// TIA Portal project "Mel7_new" (V15.1)

(* hardware
DEVICE "Станция S7-1200_1"  S7-1200 Station
   slot 0: "Rack_0"  S7-1200 Rack  Rack  V1.0
   slot 1: "01_CPU"  CPU 1215C DC/DC/DC  6ES7 215-1AG40-0XB0  V4.2
   slot 2: "AI 8x13 бит_1"  6ES7 231-4HF32-0XB0  V2.0
   slot 3: "AI 8x13 бит_2"  6ES7 231-4HF32-0XB0  V2.0
   slot 4: "AI 8x13 бит_3"  6ES7 231-4HF32-0XB0  V2.0
   slot 5: "AI 8x13 бит_4"  6ES7 231-4HF32-0XB0  V2.0
   slot 6: "AI 8xRTD_1"  SM 1231 AI8 x RTD  6ES7 231-5PF32-0XB0  V2.0
   slot 7: "AI 8xRTD_2"  SM 1231 AI8 x RTD  6ES7 231-5PF32-0XB0  V2.0
   slot 101: "CM 1243-5"  CM 1243-5  6GK7 243-5DX30-0XE0  V1.3
DEVICE "02_HMI"  KTP1200 Basic PN
   slot 0: "02_HMI"  KTP1200 Basic PN  6AV2 123-2MB03-0AX0  15.1.0.0
   slot 1: "HMI_RT_1"  KTP1200 Basic PN  6AV2 123-2MB03-0AX0  15.1.0.0
   slot 5: "02_HMI.IE_CP_1"  PROFINET Interface  15.0.1.0
      slot 1: "PROFINET Interface_1"  PROFINET Interface
         slot 1: "Port_1"  Port
DEVICE "S7300/ET200M station_1"  S7-300 station
   slot 0: "Rail_0"  Rail  6ES7 390-1***0-0AA0
   slot 2: "Slave_1"  IM 153-2  6ES7 153-2BA10-0XB0  V6.0
   slot 4: "DI 32x24VDC_1"  DI32 x 24VDC  6ES7 321-1BL00-0AA0
   slot 5: "DO 16x24VDC/0.5A_1"  DO16 x 24VDC / 0.5A  6ES7 322-1BH01-0AA0
   slot 6: "DO 16x24VDC/0.5A_2"  DO16 x 24VDC / 0.5A  6ES7 322-1BH01-0AA0
   slot 7: "AO 8x12BIT_1"  AO8 x 12 bits  6ES7 332-5HF00-0AB0
*)

// ===== PLC "01_CPU"  CPU 1215C DC/DC/DC =====

VAR_GLOBAL   // PLC tag table "Стандартная таблица переменных"
   "System_Byte" AT %MB1 : Byte;
   "FirstScan" AT %M1.0 : Bool;
   "DiagStatusUpdate" AT %M1.1 : Bool;
   "AlwaysTRUE" AT %M1.2 : Bool;
   "AlwaysFALSE" AT %M1.3 : Bool;
   "Clock_Byte" AT %MB0 : Byte;
   "Clock_10Hz" AT %M0.0 : Bool;
   "Clock_5Hz" AT %M0.1 : Bool;
   "Clock_2.5Hz" AT %M0.2 : Bool;
   "Clock_2Hz" AT %M0.3 : Bool;
   "Clock_1.25Hz" AT %M0.4 : Bool;
   "Clock_1Hz" AT %M0.5 : Bool;
   "Clock_0.625Hz" AT %M0.6 : Bool;
   "Clock_0.5Hz" AT %M0.7 : Bool;
END_VAR

TYPE "AI_STR"
   STRUCT
      "Кнопка: Закрыть фейсплату" : Bool;
      "Кнопка: Активировать HH" : Bool;   // Активация уставки НН
      "Кнопка: Активировать H" : Bool;   // Активация уставки Н
      "Кнопка: Активировать L" : Bool;   // Активация уставки L
      "Кнопка: Активировать LL" : Bool;   // Активация уставки LL
      "Кнопка: Ремонт" : Bool;   // Активация кнопки Ремонт
      Видимость : Bool;   // Видимость
      "Индикатор: Зашкал" : Bool;   // Overflow
      "Индикатор: Перелёт" : Bool;   // Overshoot range
      "Авария: Выход за HH" : Bool;   // Выход за уставку НН
      "Предупреждение: Выход за H" : Bool;   // Выход за уставку Н
      "Предупреждение: Выход за L" : Bool;   // Выход за уставку L
      "Авария: Выход за LL" : Bool;   // Выход за уставку LL
      "Индикатор: Недолет" : Bool;   // Undershoot range
      "Индикатор: Обрыв" : Bool;   // Underflow
      "Индикатор: В норме" : Bool;
      "Индикатор: HH активирована" : Bool;
      "Индикатор: H активирована" : Bool;
      "Индикатор: L активирована" : Bool;
      "Индикатор: LL активирована" : Bool;
      "Уставка: MAX" : Real := 100.0;   // Верхняя граница шкалы прибора
      "Уставка: MIN" : Real := 0.0;   // Нижняя граница шкалы прибора
      "Уставка: HH" : Real := 80.0;   // Верхняя аварийная уставка
      "Уставка: H" : Real := 70.0;   // Верхняя предупредительная уставка
      "Уставка: L" : Real := 15.0;   // Нижняя предупредительная уставка
      "Уставка: LL" : Real := 10.0;   // Нижняя аварийная уставка
      "Уставка: Перелёт" : Real := 20.0;   // Overshoot
      "Уставка: Недолёт" : Real := 4.0;   // Undershoot
      PV : Real;   // Переменная процесса
      Ток : Real;   // Токовый сигнал мА
      AnimCode : Int;
      Error : Word;   // Регистр функции ошибки
      Bipolar : Bool;   // 1 - биполярный сигнал, 0 - униполярный сигнал
      Overshoot_MIN : Int := 27649;
      Undershoot_MAX : Int := -1;
   END_STRUCT;
END_TYPE

TYPE "Motor_S"
VERSION : 0.1
   STRUCT
      Mode : Bool;   // Режим Оператор=0 Режим Автомат=1
      OperatorStart : Bool;   // Старт в режиме оператор
      AutoStart : Bool;
      ResetAlarm : Bool;
      ResetWorkTime : Bool;   // Сброс часов работы мотора
      AnimCode : Int;
      WorkTime : DInt;   // Время работы мотора
      TimeOutAccMotor : Int;
   END_STRUCT;
END_TYPE

TYPE "PID_CONT S"
   STRUCT
      COM_RST : Bool;   // Полный рестарт
      LMNR_HS : Bool;   // Верхняя граница сигнала позиционной обратной связи
      LMNR_LS : Bool;   // Нижняя граница сигнала позиционной обратной связи
      LMNS_ON : Bool := true;   // Включение сигнала ручного воздействия
      LMNUP : Bool;   // Увеличение управляющих сигналов
      LMNDN : Bool;   // Уменьшение управляющих сигналов
      PVPER_ON : Bool;   // Включение переменной процесса периферии
      CYCLE : Time := T#1s;   // Время опроса
      SP_INT : Real;   // Внутренне значение уставки
      PV_IN : Real;   // Ввод переменной уставки
      PV_PER : Word;   // Переменная процесса от периферии
      GAIN : Real := 2.0;   // Коэффицент пропорциональности
      TI : Time := T#20s;   // Время интегрирования
      DEADB_W : Real := 1.0;   // Ширина зоны нечувствительности
      PV_FAC : Real := 1.0;   // Коээфицент переменной процесса
      PV_OFF : Real;   // Смещение переменной процесса
      PULSE_TM : Time := T#3s;   // Минимальная длительность импульса
      BREAK_TM : Time := T#3s;   // Минимальная время пауза
      MTR_TM : Time := T#30s;   // Время прогона привода
      DISV : Real;   // Возмущающее воздействие
      QLMNUP : Bool;   // Увеличение управляющего сигнала
      QLMNDN : Bool;   // Уменьшение управляющего сигнала
      PV : Real;   // Переменная процесса
      ER : Real;   // Сигнал ошибки
   END_STRUCT;
END_TYPE

TYPE "DI_STR"
   STRUCT
      "BOOL" : Bool;
      "INT" : Int;
   END_STRUCT;
END_TYPE

TYPE "PID_STR"
VERSION : 0.1
   STRUCT
      SP : Real;
      PV : Real;
      Gain : Real := 2.0;
      Ti : Time := T#20s;
      Td : Time := T#10s;
      Tm_lag : Time := T#2s;
      Man_ON : Bool := true;
      MAN : Real;
      LMN_HI : Real := 100.0;
      LMN_LO : Real := 0.0;
      Reset : Bool;
      LMN : Real;
   END_STRUCT;
END_TYPE

TYPE "Motor_STR"
VERSION : 0.1
   STRUCT
      AnimCodeMotor : Int;   // Код анимации мотора
      AnimCodeKey : Int;   // Код анимации ключа: =0 Сблокированный,=1 Ручной =10,11-Ошибочная сигнализация
      TimeOutPreMotor : Int := 4;   // Таймер на нарушения мотора уставка
      TimeOutAccMotor : Int;   // Таймер на нарушения мотора аккомулятор
      TimeOutPreKey : Int := 2;   // Таймер на нарушение положения ключа уставка
      TimeOutACCKey : Int;   // Таймер на нарушение положения ключа аккомулятор
      Mode : Int;   // Режим Оператор=0 Режим Автомат=1
      PouseBeetwenON : Word;   // Пауза между включениями мотора
      WorkTime : DInt;   // Время работы мотора
      OperatorStart : Bool;   // Старт в режиме оператор
      ResetAlr : Bool;   // Сброс нарушений
      ResetWorkTime : Bool;   // Сброс часов работы мотора
      Start : Bool;   // Старт Мотора
      StartPulse : Bool;   // Старт Мотора пульс
      ModeBool : Bool;
   END_STRUCT;
END_TYPE

TYPE "Narabotki"
   STRUCT
      Hour : DInt;
      Minute : Int;
      Second : Int;
      old : Bool;
      reset : Bool;
   END_STRUCT;
END_TYPE

TYPE "Valve_STR"
VERSION : 0.1
   STRUCT
      AnimCodeValve : Int;   // Код анимации крана: =0 Нейтр,=1 Открыт, =3 закрыт, >10 Нарушения
      AnimCodeKey : Int;   // Код анимации ключа: =0 Сблокированный,=1 Ручной =10,11-Ошибочная сигнализация
      TimeOutPreValve : Int := 60;   // Таймер на нарушения движения уставка
      TimeOutAccValve : Int;   // Таймер на нарушения мотора аккомулятор
      TimeOutPreKey : Int := 2;   // Таймер на нарушение положения ключа уставка
      TimeOutACCKey : Int;   // Таймер на нарушение положения ключа аккомулятор
      Mode : Int;   // Режим Оператор=0 Режим Автомат=1
      PouseBeetwenON : Word := 16#0;   // Пауза между включениями мотора
      WorkTime : DInt;   // Время работы мотора
      OperatorOpen : Bool;   // Открытие в режиме опреатор
      OperatorClose : Bool;   // Закрытие в режиме опреатор
      ResetAlr : Bool;   // Сброс нарушений
      ResetWorkTime : Bool;   // Сброс часов работы крана
      CmdOpen : Bool;   // Команда на открытие
      CmdOpenPulse : Bool;   // Команда на открытие пульс
      CmdClose : Bool;   // Команда на закрытие
      CmdClosePulse : Bool;   // Команда на закрытие пульс
   END_STRUCT;
END_TYPE

DATA_BLOCK "01_DB_AI"   // DB1
{ S7_Optimized_Access := 'FALSE' }
VERSION : 0.1
   VAR
      L_1c : "AI_STR";
      L_1c_1 : "AI_STR";
      L_1c_2 : "AI_STR";
      L_1c_3 : "AI_STR";
      L_1c_4 : "AI_STR";
      L_1c_5 : "AI_STR";
      L_1c_6 : "AI_STR";
      L_1c_7 : "AI_STR";
      L_1c_8 : "AI_STR";
      L_1c_9 : "AI_STR";
      L_1c_10 : "AI_STR";
      L_1c_11 : "AI_STR";
      L_1c_12 : "AI_STR";
      L_1c_13 : "AI_STR";
      L_1c_14 : "AI_STR";
      L_1c_15 : "AI_STR";
      L_1c_16 : "AI_STR";
      L_1c_17 : "AI_STR";
      L_1c_18 : "AI_STR";
      L_1c_19 : "AI_STR";
      L_1c_20 : "AI_STR";
      L_1c_21 : "AI_STR";
      L_1c_22 : "AI_STR";
      L_1c_23 : "AI_STR";
      L_1c_24 : "AI_STR";
      L_1c_25 : "AI_STR";
      L_1c_26 : "AI_STR";
      L_1c_27 : "AI_STR";
      L_1c_28 : "AI_STR";
      L_1c_29 : "AI_STR";
      L_1c_30 : "AI_STR";
      L_1c_31 : "AI_STR";
      L_1c_32 : "AI_STR";
      L_1c_33 : "AI_STR";
      L_1c_36 : "AI_STR";
      L_1c_37 : "AI_STR";
      L_1c_38 : "AI_STR";
      L_1c_39 : "AI_STR";
      L_1c_40 : "AI_STR";
      L_1c_41 : "AI_STR";
      L_1c_42 : "AI_STR";
      L_1c_43 : "AI_STR";
      L_1c_44 : "AI_STR";
      L_1c_45 : "AI_STR";   // Расход руды tarir
   END_VAR
BEGIN
   L_1c_20."Кнопка: Активировать HH" := TRUE;
   L_1c_26."Кнопка: Активировать HH" := FALSE;
   L_1c."Кнопка: Закрыть фейсплату" := FALSE;
   L_1c."Кнопка: Активировать HH" := FALSE;
   L_1c."Кнопка: Активировать H" := FALSE;
   L_1c."Кнопка: Активировать L" := FALSE;
   L_1c."Кнопка: Активировать LL" := FALSE;
   L_1c."Кнопка: Ремонт" := FALSE;
   L_1c.Видимость := FALSE;
   L_1c."Индикатор: Зашкал" := FALSE;
   L_1c."Индикатор: Перелёт" := FALSE;
   L_1c."Авария: Выход за HH" := FALSE;
   L_1c."Предупреждение: Выход за H" := FALSE;
   L_1c."Предупреждение: Выход за L" := FALSE;
   L_1c."Авария: Выход за LL" := FALSE;
   L_1c."Индикатор: Недолет" := FALSE;
   L_1c."Индикатор: Обрыв" := FALSE;
   L_1c."Индикатор: В норме" := FALSE;
   L_1c."Индикатор: HH активирована" := FALSE;
   L_1c."Индикатор: H активирована" := FALSE;
   L_1c."Индикатор: L активирована" := FALSE;
   L_1c."Индикатор: LL активирована" := FALSE;
   L_1c."Уставка: MAX" := 100.0;
   L_1c."Уставка: MIN" := 0.0;
   L_1c."Уставка: HH" := 80.0;
   L_1c."Уставка: H" := 70.0;
   L_1c."Уставка: L" := 15.0;
   L_1c."Уставка: LL" := 10.0;
   L_1c."Уставка: Перелёт" := 20.0;
   L_1c."Уставка: Недолёт" := 4.0;
   L_1c.PV := 3.204572;
   L_1c.Ток := 4.512732;
   L_1c.AnimCode := 0;
   L_1c.Error := 16#0000;
   L_1c.Bipolar := FALSE;
   L_1c.Overshoot_MIN := 27649;
   L_1c.Undershoot_MAX := -1;
   L_1c_1."Кнопка: Закрыть фейсплату" := FALSE;
   L_1c_1."Кнопка: Активировать HH" := FALSE;
   L_1c_1."Кнопка: Активировать H" := FALSE;
   L_1c_1."Кнопка: Активировать L" := FALSE;
   L_1c_1."Кнопка: Активировать LL" := FALSE;
   L_1c_1."Кнопка: Ремонт" := FALSE;
   L_1c_1.Видимость := FALSE;
   L_1c_1."Индикатор: Зашкал" := FALSE;
   L_1c_1."Индикатор: Перелёт" := FALSE;
   L_1c_1."Авария: Выход за HH" := FALSE;
   L_1c_1."Предупреждение: Выход за H" := FALSE;
   L_1c_1."Предупреждение: Выход за L" := FALSE;
   L_1c_1."Авария: Выход за LL" := FALSE;
   L_1c_1."Индикатор: Недолет" := FALSE;
   L_1c_1."Индикатор: Обрыв" := FALSE;
   L_1c_1."Индикатор: В норме" := FALSE;
   L_1c_1."Индикатор: HH активирована" := FALSE;
   L_1c_1."Индикатор: H активирована" := FALSE;
   L_1c_1."Индикатор: L активирована" := FALSE;
   L_1c_1."Индикатор: LL активирована" := FALSE;
   L_1c_1."Уставка: MAX" := 100.0;
   L_1c_1."Уставка: MIN" := 0.0;
   L_1c_1."Уставка: HH" := 80.0;
   L_1c_1."Уставка: H" := 70.0;
   L_1c_1."Уставка: L" := 15.0;
   L_1c_1."Уставка: LL" := 10.0;
   L_1c_1."Уставка: Перелёт" := 20.0;
   L_1c_1."Уставка: Недолёт" := 4.0;
   L_1c_1.PV := 13.17636;
   L_1c_1.Ток := 6.108218;
   L_1c_1.AnimCode := 0;
   L_1c_1.Error := 16#0000;
   L_1c_1.Bipolar := FALSE;
   L_1c_1.Overshoot_MIN := 27649;
   L_1c_1.Undershoot_MAX := -1;
   L_1c_2."Кнопка: Закрыть фейсплату" := FALSE;
   L_1c_2."Кнопка: Активировать HH" := FALSE;
   L_1c_2."Кнопка: Активировать H" := FALSE;
   L_1c_2."Кнопка: Активировать L" := FALSE;
   L_1c_2."Кнопка: Активировать LL" := FALSE;
   L_1c_2."Кнопка: Ремонт" := FALSE;
   L_1c_2.Видимость := FALSE;
   L_1c_2."Индикатор: Зашкал" := FALSE;
   L_1c_2."Индикатор: Перелёт" := FALSE;
   L_1c_2."Авария: Выход за HH" := FALSE;
   L_1c_2."Предупреждение: Выход за H" := FALSE;
   L_1c_2."Предупреждение: Выход за L" := FALSE;
   L_1c_2."Авария: Выход за LL" := FALSE;
   L_1c_2."Индикатор: Недолет" := FALSE;
   L_1c_2."Индикатор: Обрыв" := FALSE;
   L_1c_2."Индикатор: В норме" := FALSE;
   L_1c_2."Индикатор: HH активирована" := FALSE;
   L_1c_2."Индикатор: H активирована" := FALSE;
   L_1c_2."Индикатор: L активирована" := FALSE;
   L_1c_2."Индикатор: LL активирована" := FALSE;
   L_1c_2."Уставка: MAX" := 100.0;
   L_1c_2."Уставка: MIN" := 0.0;
   L_1c_2."Уставка: HH" := 90.0;
   L_1c_2."Уставка: H" := 70.0;
   L_1c_2."Уставка: L" := 15.0;
   L_1c_2."Уставка: LL" := 10.0;
   L_1c_2."Уставка: Перелёт" := 20.0;
   L_1c_2."Уставка: Недолёт" := 4.0;
   L_1c_2.PV := 69.30339;
   L_1c_2.Ток := 15.08854;
   L_1c_2.AnimCode := 0;
   L_1c_2.Error := 16#0000;
   L_1c_2.Bipolar := FALSE;
   L_1c_2.Overshoot_MIN := 27649;
   L_1c_2.Undershoot_MAX := -1;
   L_1c_3."Кнопка: Закрыть фейсплату" := FALSE;
   L_1c_3."Кнопка: Активировать HH" := FALSE;
   L_1c_3."Кнопка: Активировать H" := FALSE;
   L_1c_3."Кнопка: Активировать L" := FALSE;
   L_1c_3."Кнопка: Активировать LL" := FALSE;
   L_1c_3."Кнопка: Ремонт" := FALSE;
   L_1c_3.Видимость := FALSE;
   L_1c_3."Индикатор: Зашкал" := FALSE;
   L_1c_3."Индикатор: Перелёт" := FALSE;
   L_1c_3."Авария: Выход за HH" := FALSE;
   L_1c_3."Предупреждение: Выход за H" := FALSE;
   L_1c_3."Предупреждение: Выход за L" := FALSE;
   L_1c_3."Авария: Выход за LL" := FALSE;
   L_1c_3."Индикатор: Недолет" := FALSE;
   L_1c_3."Индикатор: Обрыв" := FALSE;
   L_1c_3."Индикатор: В норме" := FALSE;
   L_1c_3."Индикатор: HH активирована" := FALSE;
   L_1c_3."Индикатор: H активирована" := FALSE;
   L_1c_3."Индикатор: L активирована" := FALSE;
   L_1c_3."Индикатор: LL активирована" := FALSE;
   L_1c_3."Уставка: MAX" := 100.0;
   L_1c_3."Уставка: MIN" := 0.0;
   L_1c_3."Уставка: HH" := 80.0;
   L_1c_3."Уставка: H" := 70.0;
   L_1c_3."Уставка: L" := 15.0;
   L_1c_3."Уставка: LL" := 10.0;
   L_1c_3."Уставка: Перелёт" := 20.0;
   L_1c_3."Уставка: Недолёт" := 4.0;
   L_1c_3.PV := 7.895689;
   L_1c_3.Ток := 5.26331;
   L_1c_3.AnimCode := 0;
   L_1c_3.Error := 16#0000;
   L_1c_3.Bipolar := FALSE;
   L_1c_3.Overshoot_MIN := 27649;
   L_1c_3.Undershoot_MAX := -1;
   L_1c_4."Кнопка: Закрыть фейсплату" := FALSE;
   L_1c_4."Кнопка: Активировать HH" := FALSE;
   L_1c_4."Кнопка: Активировать H" := FALSE;
   L_1c_4."Кнопка: Активировать L" := FALSE;
   L_1c_4."Кнопка: Активировать LL" := FALSE;
   L_1c_4."Кнопка: Ремонт" := FALSE;
   L_1c_4.Видимость := FALSE;
   L_1c_4."Индикатор: Зашкал" := FALSE;
   L_1c_4."Индикатор: Перелёт" := FALSE;
   L_1c_4."Авария: Выход за HH" := FALSE;
   L_1c_4."Предупреждение: Выход за H" := FALSE;
   L_1c_4."Предупреждение: Выход за L" := FALSE;
   L_1c_4."Авария: Выход за LL" := FALSE;
   L_1c_4."Индикатор: Недолет" := FALSE;
   L_1c_4."Индикатор: Обрыв" := FALSE;
   L_1c_4."Индикатор: В норме" := FALSE;
   L_1c_4."Индикатор: HH активирована" := FALSE;
   L_1c_4."Индикатор: H активирована" := FALSE;
   L_1c_4."Индикатор: L активирована" := FALSE;
   L_1c_4."Индикатор: LL активирована" := FALSE;
   L_1c_4."Уставка: MAX" := 20.0;
   L_1c_4."Уставка: MIN" := 0.0;
   L_1c_4."Уставка: HH" := 80.0;
   L_1c_4."Уставка: H" := 70.0;
   L_1c_4."Уставка: L" := 15.0;
   L_1c_4."Уставка: LL" := 10.0;
   L_1c_4."Уставка: Перелёт" := 20.0;
   L_1c_4."Уставка: Недолёт" := 4.0;
   L_1c_4.PV := 0.004340278;
   L_1c_4.Ток := 4.003472;
   L_1c_4.AnimCode := 0;
   L_1c_4.Error := 16#0000;
   L_1c_4.Bipolar := FALSE;
   L_1c_4.Overshoot_MIN := 27649;
   L_1c_4.Undershoot_MAX := -1;
   L_1c_5."Кнопка: Закрыть фейсплату" := FALSE;
   L_1c_5."Кнопка: Активировать HH" := FALSE;
   L_1c_5."Кнопка: Активировать H" := FALSE;
   L_1c_5."Кнопка: Активировать L" := FALSE;
   L_1c_5."Кнопка: Активировать LL" := FALSE;
   L_1c_5."Кнопка: Ремонт" := FALSE;
   L_1c_5.Видимость := FALSE;
   L_1c_5."Индикатор: Зашкал" := FALSE;
   L_1c_5."Индикатор: Перелёт" := FALSE;
   L_1c_5."Авария: Выход за HH" := FALSE;
   L_1c_5."Предупреждение: Выход за H" := FALSE;
   L_1c_5."Предупреждение: Выход за L" := FALSE;
   L_1c_5."Авария: Выход за LL" := FALSE;
   L_1c_5."Индикатор: Недолет" := FALSE;
   L_1c_5."Индикатор: Обрыв" := FALSE;
   L_1c_5."Индикатор: В норме" := FALSE;
   L_1c_5."Индикатор: HH активирована" := FALSE;
   L_1c_5."Индикатор: H активирована" := FALSE;
   L_1c_5."Индикатор: L активирована" := FALSE;
   L_1c_5."Индикатор: LL активирована" := FALSE;
   L_1c_5."Уставка: MAX" := 20.0;
   L_1c_5."Уставка: MIN" := 0.0;
   L_1c_5."Уставка: HH" := 80.0;
   L_1c_5."Уставка: H" := 70.0;
   L_1c_5."Уставка: L" := 15.0;
   L_1c_5."Уставка: LL" := 10.0;
   L_1c_5."Уставка: Перелёт" := 20.0;
   L_1c_5."Уставка: Недолёт" := 4.0;
   L_1c_5.PV := 0.2235243;
   L_1c_5.Ток := 4.17882;
   L_1c_5.AnimCode := 0;
   L_1c_5.Error := 16#0000;
   L_1c_5.Bipolar := FALSE;
   L_1c_5.Overshoot_MIN := 27649;
   L_1c_5.Undershoot_MAX := -1;
   L_1c_6."Кнопка: Закрыть фейсплату" := FALSE;
   L_1c_6."Кнопка: Активировать HH" := FALSE;
   L_1c_6."Кнопка: Активировать H" := FALSE;
   L_1c_6."Кнопка: Активировать L" := FALSE;
   L_1c_6."Кнопка: Активировать LL" := FALSE;
   L_1c_6."Кнопка: Ремонт" := FALSE;
   L_1c_6.Видимость := FALSE;
   L_1c_6."Индикатор: Зашкал" := FALSE;
   L_1c_6."Индикатор: Перелёт" := FALSE;
   L_1c_6."Авария: Выход за HH" := FALSE;
   L_1c_6."Предупреждение: Выход за H" := FALSE;
   L_1c_6."Предупреждение: Выход за L" := FALSE;
   L_1c_6."Авария: Выход за LL" := FALSE;
   L_1c_6."Индикатор: Недолет" := FALSE;
   L_1c_6."Индикатор: Обрыв" := FALSE;
   L_1c_6."Индикатор: В норме" := FALSE;
   L_1c_6."Индикатор: HH активирована" := FALSE;
   L_1c_6."Индикатор: H активирована" := FALSE;
   L_1c_6."Индикатор: L активирована" := FALSE;
   L_1c_6."Индикатор: LL активирована" := FALSE;
   L_1c_6."Уставка: MAX" := 1000.0;
   L_1c_6."Уставка: MIN" := 0.0;
   L_1c_6."Уставка: HH" := 80.0;
   L_1c_6."Уставка: H" := 70.0;
   L_1c_6."Уставка: L" := 15.0;
   L_1c_6."Уставка: LL" := 10.0;
   L_1c_6."Уставка: Перелёт" := 20.0;
   L_1c_6."Уставка: Недолёт" := 4.0;
   L_1c_6.PV := 0.0;
   L_1c_6.Ток := 4.0;
   L_1c_6.AnimCode := 0;
   L_1c_6.Error := 16#0000;
   L_1c_6.Bipolar := FALSE;
   L_1c_6.Overshoot_MIN := 27649;
   L_1c_6.Undershoot_MAX := -1;
   L_1c_7."Кнопка: Закрыть фейсплату" := FALSE;
   L_1c_7."Кнопка: Активировать HH" := FALSE;
   L_1c_7."Кнопка: Активировать H" := FALSE;
   L_1c_7."Кнопка: Активировать L" := FALSE;
   L_1c_7."Кнопка: Активировать LL" := FALSE;
   L_1c_7."Кнопка: Ремонт" := FALSE;
   L_1c_7.Видимость := FALSE;
   L_1c_7."Индикатор: Зашкал" := FALSE;
   L_1c_7."Индикатор: Перелёт" := FALSE;
   L_1c_7."Авария: Выход за HH" := FALSE;
   L_1c_7."Предупреждение: Выход за H" := FALSE;
   L_1c_7."Предупреждение: Выход за L" := FALSE;
   L_1c_7."Авария: Выход за LL" := FALSE;
   L_1c_7."Индикатор: Недолет" := FALSE;
   L_1c_7."Индикатор: Обрыв" := FALSE;
   L_1c_7."Индикатор: В норме" := FALSE;
   L_1c_7."Индикатор: HH активирована" := FALSE;
   L_1c_7."Индикатор: H активирована" := FALSE;
   L_1c_7."Индикатор: L активирована" := FALSE;
   L_1c_7."Индикатор: LL активирована" := FALSE;
   L_1c_7."Уставка: MAX" := 100.0;
   L_1c_7."Уставка: MIN" := 0.0;
   L_1c_7."Уставка: HH" := 80.0;
   L_1c_7."Уставка: H" := 70.0;
   L_1c_7."Уставка: L" := 15.0;
   L_1c_7."Уставка: LL" := 10.0;
   L_1c_7."Уставка: Перелёт" := 20.0;
   L_1c_7."Уставка: Недолёт" := 4.0;
   L_1c_7.PV := 0.0;
   L_1c_7.Ток := 4.0;
   L_1c_7.AnimCode := 0;
   L_1c_7.Error := 16#0000;
   L_1c_7.Bipolar := FALSE;
   L_1c_7.Overshoot_MIN := 27649;
   L_1c_7.Undershoot_MAX := -1;
   L_1c_8."Кнопка: Закрыть фейсплату" := FALSE;
   L_1c_8."Кнопка: Активировать HH" := FALSE;
   L_1c_8."Кнопка: Активировать H" := FALSE;
   L_1c_8."Кнопка: Активировать L" := FALSE;
   L_1c_8."Кнопка: Активировать LL" := FALSE;
   L_1c_8."Кнопка: Ремонт" := FALSE;
   L_1c_8.Видимость := FALSE;
   L_1c_8."Индикатор: Зашкал" := FALSE;
   L_1c_8."Индикатор: Перелёт" := FALSE;
   L_1c_8."Авария: Выход за HH" := FALSE;
   L_1c_8."Предупреждение: Выход за H" := FALSE;
   L_1c_8."Предупреждение: Выход за L" := FALSE;
   L_1c_8."Авария: Выход за LL" := FALSE;
   L_1c_8."Индикатор: Недолет" := TRUE;
   L_1c_8."Индикатор: Обрыв" := FALSE;
   L_1c_8."Индикатор: В норме" := FALSE;
   L_1c_8."Индикатор: HH активирована" := FALSE;
   L_1c_8."Индикатор: H активирована" := FALSE;
   L_1c_8."Индикатор: L активирована" := FALSE;
   L_1c_8."Индикатор: LL активирована" := FALSE;
   L_1c_8."Уставка: MAX" := 100.0;
   L_1c_8."Уставка: MIN" := 0.0;
   L_1c_8."Уставка: HH" := 80.0;
   L_1c_8."Уставка: H" := 70.0;
   L_1c_8."Уставка: L" := 15.0;
   L_1c_8."Уставка: LL" := 10.0;
   L_1c_8."Уставка: Перелёт" := 20.0;
   L_1c_8."Уставка: Недолёт" := 4.0;
   L_1c_8.PV := -0.003616898;
   L_1c_8.Ток := 3.999421;
   L_1c_8.AnimCode := 2;
   L_1c_8.Error := 16#0000;
   L_1c_8.Bipolar := FALSE;
   L_1c_8.Overshoot_MIN := 27649;
   L_1c_8.Undershoot_MAX := -1;
   L_1c_9."Кнопка: Закрыть фейсплату" := FALSE;
   L_1c_9."Кнопка: Активировать HH" := FALSE;
   L_1c_9."Кнопка: Активировать H" := FALSE;
   L_1c_9."Кнопка: Активировать L" := FALSE;
   L_1c_9."Кнопка: Активировать LL" := FALSE;
   L_1c_9."Кнопка: Ремонт" := FALSE;
   L_1c_9.Видимость := FALSE;
   L_1c_9."Индикатор: Зашкал" := FALSE;
   L_1c_9."Индикатор: Перелёт" := FALSE;
   L_1c_9."Авария: Выход за HH" := FALSE;
   L_1c_9."Предупреждение: Выход за H" := FALSE;
   L_1c_9."Предупреждение: Выход за L" := FALSE;
   L_1c_9."Авария: Выход за LL" := FALSE;
   L_1c_9."Индикатор: Недолет" := FALSE;
   L_1c_9."Индикатор: Обрыв" := FALSE;
   L_1c_9."Индикатор: В норме" := FALSE;
   L_1c_9."Индикатор: HH активирована" := FALSE;
   L_1c_9."Индикатор: H активирована" := FALSE;
   L_1c_9."Индикатор: L активирована" := FALSE;
   L_1c_9."Индикатор: LL активирована" := FALSE;
   L_1c_9."Уставка: MAX" := 20.0;
   L_1c_9."Уставка: MIN" := 0.0;
   L_1c_9."Уставка: HH" := 80.0;
   L_1c_9."Уставка: H" := 70.0;
   L_1c_9."Уставка: L" := 15.0;
   L_1c_9."Уставка: LL" := 10.0;
   L_1c_9."Уставка: Перелёт" := 20.0;
   L_1c_9."Уставка: Недолёт" := 4.0;
   L_1c_9.PV := 1.388889;
   L_1c_9.Ток := 5.111111;
   L_1c_9.AnimCode := 0;
   L_1c_9.Error := 16#0000;
   L_1c_9.Bipolar := FALSE;
   L_1c_9.Overshoot_MIN := 27649;
   L_1c_9.Undershoot_MAX := -1;
   L_1c_10."Кнопка: Закрыть фейсплату" := FALSE;
   L_1c_10."Кнопка: Активировать HH" := FALSE;
   L_1c_10."Кнопка: Активировать H" := FALSE;
   L_1c_10."Кнопка: Активировать L" := FALSE;
   L_1c_10."Кнопка: Активировать LL" := FALSE;
   L_1c_10."Кнопка: Ремонт" := FALSE;
   L_1c_10.Видимость := FALSE;
   L_1c_10."Индикатор: Зашкал" := FALSE;
   L_1c_10."Индикатор: Перелёт" := FALSE;
   L_1c_10."Авария: Выход за HH" := FALSE;
   L_1c_10."Предупреждение: Выход за H" := FALSE;
   L_1c_10."Предупреждение: Выход за L" := FALSE;
   L_1c_10."Авария: Выход за LL" := FALSE;
   L_1c_10."Индикатор: Недолет" := FALSE;
   L_1c_10."Индикатор: Обрыв" := FALSE;
   L_1c_10."Индикатор: В норме" := FALSE;
   L_1c_10."Индикатор: HH активирована" := FALSE;
   L_1c_10."Индикатор: H активирована" := FALSE;
   L_1c_10."Индикатор: L активирована" := FALSE;
   L_1c_10."Индикатор: LL активирована" := FALSE;
   L_1c_10."Уставка: MAX" := 18.0;
   L_1c_10."Уставка: MIN" := 0.0;
   L_1c_10."Уставка: HH" := 80.0;
   L_1c_10."Уставка: H" := 70.0;
   L_1c_10."Уставка: L" := 3.5;
   L_1c_10."Уставка: LL" := 3.0;
   L_1c_10."Уставка: Перелёт" := 20.0;
   L_1c_10."Уставка: Недолёт" := 4.0;
   L_1c_10.PV := 0.009765625;
   L_1c_10.Ток := 4.00868;
   L_1c_10.AnimCode := 0;
   L_1c_10.Error := 16#0000;
   L_1c_10.Bipolar := FALSE;
   L_1c_10.Overshoot_MIN := 27649;
   L_1c_10.Undershoot_MAX := -1;
   L_1c_11."Кнопка: Закрыть фейсплату" := FALSE;
   L_1c_11."Кнопка: Активировать HH" := FALSE;
   L_1c_11."Кнопка: Активировать H" := FALSE;
   L_1c_11."Кнопка: Активировать L" := FALSE;
   L_1c_11."Кнопка: Активировать LL" := FALSE;
   L_1c_11."Кнопка: Ремонт" := FALSE;
   L_1c_11.Видимость := FALSE;
   L_1c_11."Индикатор: Зашкал" := FALSE;
   L_1c_11."Индикатор: Перелёт" := FALSE;
   L_1c_11."Авария: Выход за HH" := FALSE;
   L_1c_11."Предупреждение: Выход за H" := FALSE;
   L_1c_11."Предупреждение: Выход за L" := FALSE;
   L_1c_11."Авария: Выход за LL" := FALSE;
   L_1c_11."Индикатор: Недолет" := FALSE;
   L_1c_11."Индикатор: Обрыв" := FALSE;
   L_1c_11."Индикатор: В норме" := FALSE;
   L_1c_11."Индикатор: HH активирована" := FALSE;
   L_1c_11."Индикатор: H активирована" := FALSE;
   L_1c_11."Индикатор: L активирована" := FALSE;
   L_1c_11."Индикатор: LL активирована" := FALSE;
   L_1c_11."Уставка: MAX" := 1000.0;
   L_1c_11."Уставка: MIN" := 70.0;
   L_1c_11."Уставка: HH" := 80.0;
   L_1c_11."Уставка: H" := 70.0;
   L_1c_11."Уставка: L" := 15.0;
   L_1c_11."Уставка: LL" := 10.0;
   L_1c_11."Уставка: Перелёт" := 20.0;
   L_1c_11."Уставка: Недолёт" := 4.0;
   L_1c_11.PV := 70.23546;
   L_1c_11.Ток := 4.004051;
   L_1c_11.AnimCode := 0;
   L_1c_11.Error := 16#0000;
   L_1c_11.Bipolar := FALSE;
   L_1c_11.Overshoot_MIN := 27649;
   L_1c_11.Undershoot_MAX := -1;
   L_1c_12."Кнопка: Закрыть фейсплату" := FALSE;
   L_1c_12."Кнопка: Активировать HH" := FALSE;
   L_1c_12."Кнопка: Активировать H" := FALSE;
   L_1c_12."Кнопка: Активировать L" := FALSE;
   L_1c_12."Кнопка: Активировать LL" := FALSE;
   L_1c_12."Кнопка: Ремонт" := FALSE;
   L_1c_12.Видимость := FALSE;
   L_1c_12."Индикатор: Зашкал" := FALSE;
   L_1c_12."Индикатор: Перелёт" := FALSE;
   L_1c_12."Авария: Выход за HH" := FALSE;
   L_1c_12."Предупреждение: Выход за H" := FALSE;
   L_1c_12."Предупреждение: Выход за L" := FALSE;
   L_1c_12."Авария: Выход за LL" := FALSE;
   L_1c_12."Индикатор: Недолет" := TRUE;
   L_1c_12."Индикатор: Обрыв" := FALSE;
   L_1c_12."Индикатор: В норме" := FALSE;
   L_1c_12."Индикатор: HH активирована" := FALSE;
   L_1c_12."Индикатор: H активирована" := FALSE;
   L_1c_12."Индикатор: L активирована" := FALSE;
   L_1c_12."Индикатор: LL активирована" := FALSE;
   L_1c_12."Уставка: MAX" := 250.0;
   L_1c_12."Уставка: MIN" := 0.0;
   L_1c_12."Уставка: HH" := 80.0;
   L_1c_12."Уставка: H" := 70.0;
   L_1c_12."Уставка: L" := 15.0;
   L_1c_12."Уставка: LL" := 10.0;
   L_1c_12."Уставка: Перелёт" := 20.0;
   L_1c_12."Уставка: Недолёт" := 4.0;
   L_1c_12.PV := -1.85366;
   L_1c_12.Ток := 3.881366;
   L_1c_12.AnimCode := 2;
   L_1c_12.Error := 16#0000;
   L_1c_12.Bipolar := FALSE;
   L_1c_12.Overshoot_MIN := 27649;
   L_1c_12.Undershoot_MAX := -1;
   L_1c_13."Кнопка: Закрыть фейсплату" := FALSE;
   L_1c_13."Кнопка: Активировать HH" := FALSE;
   L_1c_13."Кнопка: Активировать H" := FALSE;
   L_1c_13."Кнопка: Активировать L" := FALSE;
   L_1c_13."Кнопка: Активировать LL" := FALSE;
   L_1c_13."Кнопка: Ремонт" := FALSE;
   L_1c_13.Видимость := FALSE;
   L_1c_13."Индикатор: Зашкал" := FALSE;
   L_1c_13."Индикатор: Перелёт" := FALSE;
   L_1c_13."Авария: Выход за HH" := FALSE;
   L_1c_13."Предупреждение: Выход за H" := FALSE;
   L_1c_13."Предупреждение: Выход за L" := FALSE;
   L_1c_13."Авария: Выход за LL" := FALSE;
   L_1c_13."Индикатор: Недолет" := TRUE;
   L_1c_13."Индикатор: Обрыв" := FALSE;
   L_1c_13."Индикатор: В норме" := FALSE;
   L_1c_13."Индикатор: HH активирована" := FALSE;
   L_1c_13."Индикатор: H активирована" := FALSE;
   L_1c_13."Индикатор: L активирована" := FALSE;
   L_1c_13."Индикатор: LL активирована" := FALSE;
   L_1c_13."Уставка: MAX" := 250.0;
   L_1c_13."Уставка: MIN" := 0.0;
   L_1c_13."Уставка: HH" := 80.0;
   L_1c_13."Уставка: H" := 70.0;
   L_1c_13."Уставка: L" := 15.0;
   L_1c_13."Уставка: LL" := 10.0;
   L_1c_13."Уставка: Перелёт" := 20.0;
   L_1c_13."Уставка: Недолёт" := 4.0;
   L_1c_13.PV := -0.587746;
   L_1c_13.Ток := 3.962384;
   L_1c_13.AnimCode := 2;
   L_1c_13.Error := 16#0000;
   L_1c_13.Bipolar := FALSE;
   L_1c_13.Overshoot_MIN := 27649;
   L_1c_13.Undershoot_MAX := -1;
   L_1c_14."Кнопка: Закрыть фейсплату" := FALSE;
   L_1c_14."Кнопка: Активировать HH" := FALSE;
   L_1c_14."Кнопка: Активировать H" := FALSE;
   L_1c_14."Кнопка: Активировать L" := FALSE;
   L_1c_14."Кнопка: Активировать LL" := FALSE;
   L_1c_14."Кнопка: Ремонт" := FALSE;
   L_1c_14.Видимость := FALSE;
   L_1c_14."Индикатор: Зашкал" := FALSE;
   L_1c_14."Индикатор: Перелёт" := FALSE;
   L_1c_14."Авария: Выход за HH" := FALSE;
   L_1c_14."Предупреждение: Выход за H" := FALSE;
   L_1c_14."Предупреждение: Выход за L" := FALSE;
   L_1c_14."Авария: Выход за LL" := FALSE;
   L_1c_14."Индикатор: Недолет" := TRUE;
   L_1c_14."Индикатор: Обрыв" := FALSE;
   L_1c_14."Индикатор: В норме" := FALSE;
   L_1c_14."Индикатор: HH активирована" := FALSE;
   L_1c_14."Индикатор: H активирована" := FALSE;
   L_1c_14."Индикатор: L активирована" := FALSE;
   L_1c_14."Индикатор: LL активирована" := FALSE;
   L_1c_14."Уставка: MAX" := 250.0;
   L_1c_14."Уставка: MIN" := 0.0;
   L_1c_14."Уставка: HH" := 80.0;
   L_1c_14."Уставка: H" := 70.0;
   L_1c_14."Уставка: L" := 15.0;
   L_1c_14."Уставка: LL" := 10.0;
   L_1c_14."Уставка: Перелёт" := 20.0;
   L_1c_14."Уставка: Недолёт" := 4.0;
   L_1c_14.PV := -5.570024;
   L_1c_14.Ток := 3.643518;
   L_1c_14.AnimCode := 2;
   L_1c_14.Error := 16#0000;
   L_1c_14.Bipolar := FALSE;
   L_1c_14.Overshoot_MIN := 27649;
   L_1c_14.Undershoot_MAX := -1;
   L_1c_15."Кнопка: Закрыть фейсплату" := FALSE;
   L_1c_15."Кнопка: Активировать HH" := FALSE;
   L_1c_15."Кнопка: Активировать H" := FALSE;
   L_1c_15."Кнопка: Активировать L" := FALSE;
   L_1c_15."Кнопка: Активировать LL" := FALSE;
   L_1c_15."Кнопка: Ремонт" := FALSE;
   L_1c_15.Видимость := FALSE;
   L_1c_15."Индикатор: Зашкал" := FALSE;
   L_1c_15."Индикатор: Перелёт" := FALSE;
   L_1c_15."Авария: Выход за HH" := FALSE;
   L_1c_15."Предупреждение: Выход за H" := FALSE;
   L_1c_15."Предупреждение: Выход за L" := FALSE;
   L_1c_15."Авария: Выход за LL" := FALSE;
   L_1c_15."Индикатор: Недолет" := FALSE;
   L_1c_15."Индикатор: Обрыв" := FALSE;
   L_1c_15."Индикатор: В норме" := FALSE;
   L_1c_15."Индикатор: HH активирована" := FALSE;
   L_1c_15."Индикатор: H активирована" := TRUE;
   L_1c_15."Индикатор: L активирована" := FALSE;
   L_1c_15."Индикатор: LL активирована" := FALSE;
   L_1c_15."Уставка: MAX" := 60.0;
   L_1c_15."Уставка: MIN" := 0.0;
   L_1c_15."Уставка: HH" := 45.0;
   L_1c_15."Уставка: H" := 45.0;
   L_1c_15."Уставка: L" := 1.1;
   L_1c_15."Уставка: LL" := 1.1;
   L_1c_15."Уставка: Перелёт" := 20.0;
   L_1c_15."Уставка: Недолёт" := 4.0;
   L_1c_15.PV := 0.008680556;
   L_1c_15.Ток := 4.002315;
   L_1c_15.AnimCode := 0;
   L_1c_15.Error := 16#0000;
   L_1c_15.Bipolar := FALSE;
   L_1c_15.Overshoot_MIN := 27649;
   L_1c_15.Undershoot_MAX := -1;
   L_1c_16."Кнопка: Закрыть фейсплату" := FALSE;
   L_1c_16."Кнопка: Активировать HH" := FALSE;
   L_1c_16."Кнопка: Активировать H" := FALSE;
   L_1c_16."Кнопка: Активировать L" := FALSE;
   L_1c_16."Кнопка: Активировать LL" := FALSE;
   L_1c_16."Кнопка: Ремонт" := FALSE;
   L_1c_16.Видимость := FALSE;
   L_1c_16."Индикатор: Зашкал" := FALSE;
   L_1c_16."Индикатор: Перелёт" := FALSE;
   L_1c_16."Авария: Выход за HH" := FALSE;
   L_1c_16."Предупреждение: Выход за H" := FALSE;
   L_1c_16."Предупреждение: Выход за L" := FALSE;
   L_1c_16."Авария: Выход за LL" := FALSE;
   L_1c_16."Индикатор: Недолет" := FALSE;
   L_1c_16."Индикатор: Обрыв" := FALSE;
   L_1c_16."Индикатор: В норме" := FALSE;
   L_1c_16."Индикатор: HH активирована" := FALSE;
   L_1c_16."Индикатор: H активирована" := FALSE;
   L_1c_16."Индикатор: L активирована" := FALSE;
   L_1c_16."Индикатор: LL активирована" := FALSE;
   L_1c_16."Уставка: MAX" := 150.0;
   L_1c_16."Уставка: MIN" := 0.0;
   L_1c_16."Уставка: HH" := 65.0;
   L_1c_16."Уставка: H" := 55.0;
   L_1c_16."Уставка: L" := 15.0;
   L_1c_16."Уставка: LL" := 10.0;
   L_1c_16."Уставка: Перелёт" := 20.0;
   L_1c_16."Уставка: Недолёт" := 4.0;
   L_1c_16.PV := 23.4;
   L_1c_16.Ток := 0.0;
   L_1c_16.AnimCode := 0;
   L_1c_16.Error := 16#0000;
   L_1c_16.Bipolar := FALSE;
   L_1c_16.Overshoot_MIN := 27649;
   L_1c_16.Undershoot_MAX := -1;
   L_1c_17."Кнопка: Закрыть фейсплату" := FALSE;
   L_1c_17."Кнопка: Активировать HH" := FALSE;
   L_1c_17."Кнопка: Активировать H" := FALSE;
   L_1c_17."Кнопка: Активировать L" := FALSE;
   L_1c_17."Кнопка: Активировать LL" := FALSE;
   L_1c_17."Кнопка: Ремонт" := FALSE;
   L_1c_17.Видимость := FALSE;
   L_1c_17."Индикатор: Зашкал" := FALSE;
   L_1c_17."Индикатор: Перелёт" := FALSE;
   L_1c_17."Авария: Выход за HH" := FALSE;
   L_1c_17."Предупреждение: Выход за H" := FALSE;
   L_1c_17."Предупреждение: Выход за L" := FALSE;
   L_1c_17."Авария: Выход за LL" := FALSE;
   L_1c_17."Индикатор: Недолет" := FALSE;
   L_1c_17."Индикатор: Обрыв" := FALSE;
   L_1c_17."Индикатор: В норме" := FALSE;
   L_1c_17."Индикатор: HH активирована" := FALSE;
   L_1c_17."Индикатор: H активирована" := FALSE;
   L_1c_17."Индикатор: L активирована" := FALSE;
   L_1c_17."Индикатор: LL активирована" := FALSE;
   L_1c_17."Уставка: MAX" := 160.0;
   L_1c_17."Уставка: MIN" := 0.0;
   L_1c_17."Уставка: HH" := 80.0;
   L_1c_17."Уставка: H" := 70.0;
   L_1c_17."Уставка: L" := 15.0;
   L_1c_17."Уставка: LL" := 10.0;
   L_1c_17."Уставка: Перелёт" := 20.0;
   L_1c_17."Уставка: Недолёт" := 4.0;
   L_1c_17.PV := 0.0;
   L_1c_17.Ток := 0.0;
   L_1c_17.AnimCode := 0;
   L_1c_17.Error := 16#0000;
   L_1c_17.Bipolar := FALSE;
   L_1c_17.Overshoot_MIN := 27649;
   L_1c_17.Undershoot_MAX := -1;
   L_1c_18."Кнопка: Закрыть фейсплату" := FALSE;
   L_1c_18."Кнопка: Активировать HH" := FALSE;
   L_1c_18."Кнопка: Активировать H" := FALSE;
   L_1c_18."Кнопка: Активировать L" := FALSE;
   L_1c_18."Кнопка: Активировать LL" := FALSE;
   L_1c_18."Кнопка: Ремонт" := FALSE;
   L_1c_18.Видимость := FALSE;
   L_1c_18."Индикатор: Зашкал" := FALSE;
   L_1c_18."Индикатор: Перелёт" := FALSE;
   L_1c_18."Авария: Выход за HH" := FALSE;
   L_1c_18."Предупреждение: Выход за H" := FALSE;
   L_1c_18."Предупреждение: Выход за L" := FALSE;
   L_1c_18."Авария: Выход за LL" := FALSE;
   L_1c_18."Индикатор: Недолет" := FALSE;